(* Logix 5000 project; controller PLC_MCC1300_75F1 vendor 1 type 14 code 166 rev 32.11; software revision 32.04; part 63 of 83 *)
(* tags used below, declared in another part *)
   AUX_xInitialize : BOOL;
   CONST_rgdDestMask : DINT[32];   // Destination Mask
   CONST_tPlant : UDT_PLANT_CONSTANTS;
   GP_TrackingGetFirstPlateInConveyor : GP_TrackingGetFirstPlateInConveyor;
   GP_TrackingPresencePlate : GP_TrackingPresencePlate;
   GP_TrackingSearchPlate : GP_TrackingSearchPlate;
   M315_M1_DR_R1 : AXIS_CIP_DRIVE;
   M315_xReqStopPrevConvForPos : BOOL;
   M315Popup : MAC_Popup_ZC[2];
   M315Popup_xDrivePosEnable : BOOL;
   TMP_d : DINT;
   TMP_dIndex : DINT;
   TMP_dIndex2 : DINT;
   TMP_dIndex3 : DINT;
   TMP_dStart0 : DINT;
   TMP_dStart1 : DINT;
   TMP_dStartSearchStop : DINT;
   TMP_dStop0 : DINT;
   TMP_dStop1 : DINT;
   TMP_dStopSearchStop : DINT;
   TMP_StartPlusLength : DINT;
   TMP_xAllLiteToCullet : BOOL;
   TMP_xAtLeastOneForSideLeg : BOOL;
   TMP_xPosHead : BOOL;
   TMP_xReqStopM315M1 : BOOL;
   TMP_xReqStopM315M2 : BOOL;
   TMP_xReqStopM315M3 : BOOL;
   xAlwaysOFF : BOOL;
   xDebugOFF : BOOL;
   Z300_BufferPlate : UDT_LINE_BUFFER_PLATE;
   Z300_Conveyor : UDT_StandConv[29];
   Z300_Conveyor_IN_MOTION : MAC_Conveyor_ZC_IN_MOTION[29];
   Z300_LineTracking : UDT_LINE_TRACKING;
(* MainProgram, continued *)

   37: XIC(Z300_Conveyor[26].OUTPUT_xPositioning.0)[[XIC(Z300_Conveyor_IN_MOTION[26].DR_MAM_M[0].PC) ,XIC(xAlwaysOFF) ADD(Z300_LineTracking.rgtTrkConv[26].dStartPosition_cmm,Z300_Conveyor[26].AUX_rgdTarget_cmm[0],TMP_d) SUB(TMP_d,Z300_LineTracking.rgtTrkConv[26].dActualRamp_cmm[0],TMP_d) GEQ(Z300_BufferPlate.rgtPlate[TMP_dIndex].tTracking.dPositionHead_cmm,TMP_d) ] ,XIO(xDebugOFF) XIC(Z300_Conveyor[26].ST_xPositionReached) ][OTE(Z300_Conveyor[26].ST_xPositionReached) ,MOV(M315Popup[0].AUX_dIndexPositioning,TMP_dIndex) JSR(sbrTrackingPositioningDone,3,TMP_dIndex,TMP_xPosHead,Z300_Conveyor[26].AUX_rgdTarget_cmm[0]) ];
   38: XIC(Z300_Conveyor[27].OUTPUT_xPositioning.0)[[XIC(Z300_Conveyor_IN_MOTION[27].DR_MAM_M[0].PC) ,XIC(xAlwaysOFF) ADD(Z300_LineTracking.rgtTrkConv[26].dStartPosition_cmm,Z300_Conveyor[26].AUX_rgdTarget_cmm[0],TMP_d) SUB(TMP_d,Z300_LineTracking.rgtTrkConv[26].dActualRamp_cmm[0],TMP_d) GEQ(Z300_BufferPlate.rgtPlate[TMP_dIndex].tTracking.dPositionHead_cmm,TMP_d) ] ,XIO(xDebugOFF) XIC(Z300_Conveyor[27].ST_xPositionReached) ][OTE(Z300_Conveyor[27].ST_xPositionReached) ,MOV(M315Popup[0].AUX_dIndexPositioning,TMP_dIndex) JSR(sbrTrackingPositioningDone,3,TMP_dIndex,TMP_xPosHead,Z300_Conveyor[26].AUX_rgdTarget_cmm[0]) ];
   39: XIC(Z300_Conveyor[28].OUTPUT_xPositioning.0)[XIC(Z300_Conveyor_IN_MOTION[28].DR_MAM_M[0].PC) ,XIC(xAlwaysOFF) ADD(Z300_LineTracking.rgtTrkConv[26].dStartPosition_cmm,Z300_Conveyor[26].AUX_rgdTarget_cmm[0],TMP_d) SUB(TMP_d,Z300_LineTracking.rgtTrkConv[26].dActualRamp_cmm[0],TMP_d) GEQ(Z300_BufferPlate.rgtPlate[TMP_dIndex].tTracking.dPositionHead_cmm,TMP_d) ,XIO(xAlwaysOFF) XIC(Z300_Conveyor[28].ST_xPositionReached) ][OTE(Z300_Conveyor[28].ST_xPositionReached) ,MOV(M315Popup[0].AUX_dIndexPositioning,TMP_dIndex) JSR(sbrTrackingPositioningDone,3,TMP_dIndex,TMP_xPosHead,Z300_Conveyor[26].AUX_rgdTarget_cmm[0]) ];
   // Head positioning done
   40: [XIC(Z300_Conveyor[26].xReqPositioningHead) ,XIC(Z300_Conveyor[27].xReqPositioningHead) ,XIC(Z300_Conveyor[28].xReqPositioningHead) ][XIC(Z300_Conveyor[26].ST_xPositionReached) XIC(Z300_Conveyor[27].ST_xPositionReached) [XIC(Z300_Conveyor[28].ST_xPositionReached) ,XIO(Z300_Conveyor[28].xReqPositioningHead) ] ,XIC(Z300_Conveyor[26].xReqStop) XIO(Z300_Conveyor[26].ST_xRotationFeedback) XIC(Z300_Conveyor[27].xReqStop) XIO(Z300_Conveyor[27].ST_xRotationFeedback) [XIC(Z300_Conveyor[28].xReqStop) XIO(Z300_Conveyor[28].ST_xRotationFeedback) ,XIO(Z300_Conveyor[28].xReqPositioningHead) ] ,XIC(M315Popup[0].OS_xTimeoutPositioning) ,XIC(xDebugOFF) XIO(M315Popup[0].ST_xIndexConsPositioning) ,XIC(Z300_Conveyor[26].ST_xCleaningEnabled) ,XIC(Z300_Conveyor[26].ST_xFaulted) ,XIC(Z300_Conveyor[27].ST_xFaulted) ,XIC(Z300_Conveyor[28].ST_xFaulted) ][OTU(Z300_Conveyor[26].xReqPositioningHead) ,OTU(Z300_Conveyor[27].xReqPositioningHead) ,OTU(Z300_Conveyor[28].xReqPositioningHead) ,XIO(Z300_Conveyor[26].ST_xFaulted) XIO(Z300_Conveyor[27].ST_xFaulted) XIO(Z300_Conveyor[28].ST_xFaulted) XIO(Z300_Conveyor[26].ST_xCleaningEnabled) XIO(M315Popup[0].OS_xTimeoutPositioning) XIC(M315Popup[0].ST_xIndexConsPositioning) MOV(M315Popup[0].AUX_dIndexPositioning,TMP_dIndex) [OTL(Z300_BufferPlate.rgtPlate[TMP_dIndex].tData.tFlag.tConveyor.xDoneHeadPositioning) ,JSR(sbrTrackingPositioningDone,3,TMP_dIndex,TMP_xPosHead,Z300_Conveyor[26].AUX_rgdTarget_cmm[0]) ,MOV(M315Popup[0].AUX_dIndexPositioning,M315Popup[0].AUX_dIndexPlatePositioned) ] ,MOV(0,M315Popup[0].AUX_dIndexHead) ];
   // When plate tail has passed previous conveyor remove positioning
   41: [XIC(Z300_Conveyor[26].xReqPositioningHead) ,XIC(Z300_Conveyor[27].xReqPositioningHead) ,XIC(Z300_Conveyor[28].xReqPositioningHead) ][XIO(M315Popup[0].ST_xPrevConvFreeAfterPos) NEQ(M315Popup[0].AUX_dIndexPositioning,0) ,XIC(M315Popup[0].ST_xPrevConvFreeAfterPos) EQU(M315Popup[0].AUX_dIndexPositioning,M315Popup[0].AUX_dLastIndexFreeForPos) ][XIC(Z300_Conveyor[25].xReqPositioningHead) MOV(M315Popup[0].AUX_dIndexPositioning,TMP_dIndex) GEQ(Z300_BufferPlate.rgtPlate[TMP_dIndex].tTracking.dPositionTail_cmm,Z300_LineTracking.rgtTrkConv[25].dEndPosition_cmm) ,XIC(M315Popup[0].ST_xPrevConvFreeAfterPos) ][OTU(Z300_Conveyor[25].xReqPositioningHead) ,[XIC(Z300_Conveyor[26].ST_xRotationFeedback) ,XIC(Z300_Conveyor[26].ST_xDriveInDec) ] OTE(M315Popup[0].ST_xPrevConvFreeAfterPos) ,ONS(M315Popup[0].OS_xLastFreeForPos) MOV(M315Popup[0].AUX_dIndexPositioning,M315Popup[0].AUX_dLastIndexFreeForPos) ];
   // Tail positioning done
   42: [XIC(Z300_Conveyor[26].xReqPositioningTail) ,XIC(Z300_Conveyor[27].xReqPositioningTail) ,XIC(Z300_Conveyor[28].xReqPositioningTail) ][XIC(Z300_Conveyor[26].ST_xPositionReached) XIC(Z300_Conveyor[27].ST_xPositionReached) [XIC(Z300_Conveyor[28].ST_xPositionReached) ,XIO(Z300_Conveyor[28].xReqPositioningTail) ] ,XIC(M315Popup[0].OS_xTimeoutPositioning) ,XIO(M315Popup[0].ST_xIndexConsPositioning) ,XIC(Z300_Conveyor[26].ST_xCleaningEnabled) ,XIC(Z300_Conveyor[26].ST_xFaulted) ,XIC(Z300_Conveyor[27].ST_xFaulted) ,XIC(Z300_Conveyor[28].ST_xFaulted) ][OTU(Z300_Conveyor[26].xReqPositioningTail) ,OTU(Z300_Conveyor[27].xReqPositioningTail) ,OTU(Z300_Conveyor[28].xReqPositioningTail) ,XIO(Z300_Conveyor[26].ST_xFaulted) XIO(Z300_Conveyor[27].ST_xFaulted) XIO(Z300_Conveyor[28].ST_xFaulted) XIO(Z300_Conveyor[26].ST_xCleaningEnabled) XIO(M315Popup[0].OS_xTimeoutPositioning) MOV(M315Popup[0].AUX_tSearchPlateData.dIndex,TMP_dIndex) [OTL(Z300_BufferPlate.rgtPlate[TMP_dIndex].tData.tFlag.tConveyor.xDoneTailPositioning) ,JSR(sbrTrackingPositioningDone,3,TMP_dIndex,TMP_xPosHead,Z300_Conveyor[26].AUX_rgdTarget_cmm[0]) ,XIO(xDebugOFF) MOV(M315Popup[0].AUX_dIndexPositioning,M315Popup[0].AUX_dIndexPlatePositioned) ] ,MOV(0,M315Popup[0].AUX_dIndexTail) ];
   // Timeout positioning
   43: [[XIC(Z300_Conveyor[26].xReqPositioningHead) ,XIC(Z300_Conveyor[27].xReqPositioningHead) ,XIC(Z300_Conveyor[28].xReqPositioningHead) ] MOV(M315Popup[0].AUX_dIndexPositioning,TMP_dIndex) GEQ(Z300_BufferPlate.rgtPlate[TMP_dIndex].tTracking.dPositionHead_cmm,M315Popup[0].AUX_dPosTimeout) XIO(Z300_BufferPlate.rgtPlate[TMP_dIndex].tData.tFlag.tConveyor.xDoneHeadPositioning) ,[XIC(Z300_Conveyor[26].xReqPositioningTail) ,XIC(Z300_Conveyor[27].xReqPositioningTail) ,XIC(Z300_Conveyor[28].xReqPositioningTail) ] MOV(M315Popup[0].AUX_dIndexPositioning,TMP_dIndex) GEQ(Z300_BufferPlate.rgtPlate[TMP_dIndex].tTracking.dPositionTail_cmm,M315Popup[0].AUX_dPosTimeout) XIO(Z300_BufferPlate.rgtPlate[TMP_dIndex].tData.tFlag.tConveyor.xDoneTailPositioning) ]OTE(M315Popup[0].OS_xTimeoutPositioning);
   44: XIC(Z300_Conveyor[25].xReqPositioningHead)XIO(M315Popup[0].AUX_tSearchPlateData.xPlateHooked)OTU(Z300_Conveyor[25].xReqPositioningHead);
   45: XIC(Z300_Conveyor[25].xReqPositioningTail)XIO(M315Popup[0].AUX_tSearchPlateData.xPlateHooked)OTU(Z300_Conveyor[25].xReqPositioningTail);
   46: XIC(Z300_Conveyor[26].xReqPositioningHead)XIO(M315Popup[0].AUX_tSearchPlateData.xPlateHooked)OTU(Z300_Conveyor[26].xReqPositioningHead);
   47: XIC(Z300_Conveyor[26].xReqPositioningTail)XIO(M315Popup[0].AUX_tSearchPlateData.xPlateHooked)OTU(Z300_Conveyor[26].xReqPositioningTail);
   48: XIC(Z300_Conveyor[27].xReqPositioningHead)XIO(M315Popup[0].AUX_tSearchPlateData.xPlateHooked)OTU(Z300_Conveyor[27].xReqPositioningHead);
   49: XIC(Z300_Conveyor[27].xReqPositioningTail)XIO(M315Popup[0].AUX_tSearchPlateData.xPlateHooked)OTU(Z300_Conveyor[27].xReqPositioningTail);
   50: XIC(Z300_Conveyor[28].xReqPositioningHead)XIO(M315Popup[0].AUX_tSearchPlateData.xPlateHooked)OTU(Z300_Conveyor[28].xReqPositioningHead);
   51: XIC(Z300_Conveyor[28].xReqPositioningTail)XIO(M315Popup[0].AUX_tSearchPlateData.xPlateHooked)OTU(Z300_Conveyor[28].xReqPositioningTail);
   // #####_PRESENCE_PLATE_ON_POPUP_AFTER_POSITIONING_#####
   52: NOP();
   // Search on whole popup size
   53: ADD(0,M315Popup[0].AUX_dStartPosition_cmm,TMP_dStartSearchStop)ADD(70000,M315Popup[1].AUX_dEndPosition_cmm,TMP_dStopSearchStop)XIC(M315Popup[0].ST_xPlateToSinglePositioning)ADD(0,M315Popup[0].AUX_dStartPosition_cmm,TMP_dStartSearchStop)ADD(70000,M315Popup[0].AUX_dEndPosition_cmm,TMP_dStopSearchStop);
   54: GP_TrackingSearchPlate(GP_TrackingSearchPlate,TMP_dStopSearchStop,TMP_dStartSearchStop,0,Z300_LineTracking,M315Popup[0].tSearchPlateStop,CONST_tPlant.dNumOfConveyors,CONST_tPlant.dNumCapsConveyor,Z300_BufferPlate);
   55: XIC(M315Popup[0].tSearchPlateStop.xHeadPresence)MOV(M315Popup[0].tSearchPlateStop.rgdHeadPointer[0],M315Popup[0].AUX_dIndexPlateStop);
   56: XIO(M315Popup[0].tSearchPlateStop.xHeadPresence)XIC(M315Popup[0].tSearchPlateStop.xTailPresence)MOV(M315Popup[0].tSearchPlateStop.rgdTailPointer[0],M315Popup[0].AUX_dIndexPlateStop);
   57: [XIO(M315Popup[0].tSearchPlateStop.xHeadPresence) XIO(M315Popup[0].tSearchPlateStop.xTailPresence) ,XIC(Z300_Conveyor[26].ST_xCleaningEnabled) ]MOV(0,M315Popup[0].AUX_dIndexPlateStop);
   58: [XIC(M315Popup[0].tSearchPlateStop.xHeadPresence) ,XIC(M315Popup[0].tSearchPlateStop.xTailPresence) ][OTU(TMP_xAtLeastOneForSideLeg) ,OTL(TMP_xAllLiteToCullet) ];
   59: [XIC(M315Popup[0].tSearchPlateStop.xHeadPresence) ,XIC(M315Popup[0].tSearchPlateStop.xTailPresence) ]JSR(sbrCheckConvoyZCDestination,5,M315Popup[0].AUX_dIndexPlateStop,M315Popup[0].AUX_dDestMaskOppOpSide,CONST_rgdDestMask[24],TMP_xAtLeastOneForSideLeg,TMP_xAllLiteToCullet,TMP_xAtLeastOneForSideLeg,TMP_xAllLiteToCullet)XIC(TMP_xAtLeastOneForSideLeg)[EQU(M315Popup[0].AUX_dIndexPositioning,M315Popup[0].AUX_dIndexPlateStop) ,EQU(M315Popup[0].AUX_dIndexPlatePositioned,M315Popup[0].AUX_dIndexPlateStop) ,EQU(M315Popup[0].tSearchPlateStop.rgdHeadPointer[1],M315Popup[0].AUX_dIndexPlateStop) ,EQU(M315Popup[0].tSearchPlateStop.rgdHeadPointer[1],M315Popup[0].AUX_dIndexPlatePositioned) ,EQU(M315Popup[0].tSearchPlateStop.rgdTailPointer[1],M315Popup[0].AUX_dIndexPlateStop) ,EQU(M315Popup[0].tSearchPlateStop.rgdTailPointer[1],M315Popup[0].AUX_dIndexPlatePositioned) ,XIO(xDebugOFF) ]OTE(M315Popup[0].ST_xPlateStopToPopup);
   // IndexPlatePositioned valorizzata qui solo per la simulazione (da togliere)
   60: XIC(M315Popup[0].AUX_tSearchPlateData.xPlateHooked)[XIC(M315Popup[0].tSearchPlateStop.xHeadPresence) ,XIC(M315Popup[0].tSearchPlateStop.xTailPresence) ,XIO(M315Popup[1].ST_xPlateToSinglePositioning) EQU(M315Popup[0].AUX_dIndexPositioning,Z300_LineTracking.rgtTrkConv[26].Cap[0].dPointer) ,XIO(M315Popup[1].ST_xPlateToSinglePositioning) EQU(M315Popup[0].AUX_dIndexPlatePositioned,Z300_LineTracking.rgtTrkConv[26].Cap[0].dPointer) ][XIC(TMP_xPosHead) MOV(M315Popup[0].AUX_dIndexPositioning,TMP_dIndex) XIC(Z300_BufferPlate.rgtPlate[TMP_dIndex].tData.tFlag.tConveyor.xDoneHeadPositioning) ,XIO(TMP_xPosHead) MOV(M315Popup[0].AUX_dIndexPositioning,TMP_dIndex) XIC(Z300_BufferPlate.rgtPlate[TMP_dIndex].tData.tFlag.tConveyor.xDoneTailPositioning) ]XIO(M315Popup_xDrivePosEnable)XIC(M315Popup[0].ST_xPlateStopToPopup)[OTE(TMP_xReqStopM315M1) ,OTE(TMP_xReqStopM315M2) ,XIO(M315Popup[0].ST_xPlateToSinglePositioning) OTE(TMP_xReqStopM315M3) ];
   61: XIO(xDebugOFF)XIC(Z300_Conveyor[26].OUTPUT_xPositioning.0)OTE(Z300_Conveyor[26].xReqBypassEndStop);
   62: XIO(xDebugOFF)XIC(Z300_Conveyor[27].OUTPUT_xPositioning.0)OTE(Z300_Conveyor[27].xReqBypassEndStop);
   63: XIO(xDebugOFF)XIC(Z300_Conveyor[28].OUTPUT_xPositioning.0)OTE(Z300_Conveyor[28].xReqBypassEndStop);
   64: [XIC(TMP_xReqStopM315M1) ,XIC(M315Popup[0].PH_xDescend) ]OTE(Z300_Conveyor[26].xReqStop);
   65: [XIC(TMP_xReqStopM315M2) ,XIC(M315Popup[0].PH_xDescend) ]OTE(Z300_Conveyor[27].xReqStop);
   66: [XIC(TMP_xReqStopM315M3) ,XIC(M315Popup[1].PH_xDescend) ]OTE(Z300_Conveyor[28].xReqStop);
   // Stop tracking update while ending positioning
   67: XIO(xDebugOFF)XIC(M315Popup[0].AUX_tSearchPlateData.xPlateHooked)MOV(M315Popup[0].AUX_dIndexPositioning,TMP_dIndex)XIC(M315Popup_xDrivePosEnable)[ADD(Z300_LineTracking.rgtTrkConv[26].dStartPosition_cmm,Z300_Conveyor[26].AUX_rgdTarget_cmm[0],TMP_d) SUB(TMP_d,Z300_LineTracking.rgtTrkConv[26].dActualRamp_cmm[0],TMP_d) GEQ(Z300_BufferPlate.rgtPlate[TMP_dIndex].tTracking.dPositionHead_cmm,TMP_d) ,ADD(Z300_LineTracking.rgtTrkConv[26].dStartPosition_cmm,Z300_BufferPlate.rgtPlate[TMP_dIndex].tData.rgtCap[0].dConvTotLength_cmm,TMP_StartPlusLength) GEQ(Z300_BufferPlate.rgtPlate[TMP_dIndex].tTracking.dPositionHead_cmm,TMP_StartPlusLength) ][XIC(M315Popup[0].ST_xPlateStopToPopup) ,XIC(M315Popup[1].ST_xPlateStopToPopup) ]XIC(Z300_Conveyor_IN_MOTION[26].DR_MAM_M[0].IP)XIO(Z300_Conveyor_IN_MOTION[26].DR_MAM_M[0].PC)XIO(Z300_Conveyor_IN_MOTION[26].DR_MAM_M[0].ER)[OTE(Z300_BufferPlate.rgtPlate[TMP_dIndex].tTracking.xHoldAdvancement) ,ADD(M315Popup[0].AUX_dPosPhotocell_cmm,Z300_Conveyor[26].AUX_rgdTarget_cmm[0],TMP_d) JSR(sbrUpdateTrackingConvoyPosition,2,TMP_dIndex,TMP_d) ];
   // Stop tracking update while ending positioning
   68: XIC(M315Popup[0].AUX_tSearchPlateData.xPlateHooked)[XIC(Z300_LineTracking.rgtTrkConv[26].xGlassPresence) ,XIC(Z300_LineTracking.rgtTrkConv[27].xGlassPresence) ,XIC(Z300_LineTracking.rgtTrkConv[28].xGlassPresence) ]MOV(M315Popup[0].AUX_dIndexPositioning,TMP_dIndex)[LES(Z300_BufferPlate.rgtPlate[TMP_dIndex].tData.dTotalCaps,2) ,XIO(xDebugOFF) ]XIC(M315Popup_xDrivePosEnable)XIO(M315_M1_DR_R1.Registration1InputStatus)[ADD(Z300_LineTracking.rgtTrkConv[26].dStartPosition_cmm,Z300_Conveyor[26].AUX_rgdTarget_cmm[0],TMP_d) SUB(TMP_d,Z300_LineTracking.rgtTrkConv[26].dActualRamp_cmm[0],TMP_d) GEQ(Z300_BufferPlate.rgtPlate[TMP_dIndex].tTracking.dPositionHead_cmm,TMP_d) ,ADD(Z300_LineTracking.rgtTrkConv[26].dStartPosition_cmm,Z300_BufferPlate.rgtPlate[TMP_dIndex].tData.rgtCap[0].dConvTotLength_cmm,TMP_StartPlusLength) GEQ(Z300_BufferPlate.rgtPlate[TMP_dIndex].tTracking.dPositionHead_cmm,TMP_StartPlusLength) ]OTE(M315_xReqStopPrevConvForPos);
   69: XIO(xDebugOFF)XIC(Z300_BufferPlate.rgtPlate[TMP_dIndex].tTracking.xHoldAdvancement)GRT(Z300_BufferPlate.rgtPlate[TMP_dIndex].tTracking.dNextCapIndex,0)MOV(Z300_BufferPlate.rgtPlate[TMP_dIndex].tTracking.dNextCapIndex,TMP_dIndex2)OTE(Z300_BufferPlate.rgtPlate[TMP_dIndex2].tTracking.xHoldAdvancement);
   70: XIO(xDebugOFF)XIC(Z300_BufferPlate.rgtPlate[TMP_dIndex2].tTracking.xHoldAdvancement)GRT(Z300_BufferPlate.rgtPlate[TMP_dIndex2].tTracking.dNextCapIndex,0)MOV(Z300_BufferPlate.rgtPlate[TMP_dIndex2].tTracking.dNextCapIndex,TMP_dIndex3)OTE(Z300_BufferPlate.rgtPlate[TMP_dIndex3].tTracking.xHoldAdvancement);
   // #####_PRESENCE_PLATE_UNDER_POPUP_#####
   71: NOP();
   72: [XIC(Z300_Conveyor[25].ST_xRotationFeedback) SUB(M315Popup[0].AUX_dStartPosition_cmm,25000,TMP_dStart0) ,XIO(Z300_Conveyor[25].ST_xRotationFeedback) SUB(M315Popup[0].AUX_dStartPosition_cmm,0,TMP_dStart0) ]ADD(M315Popup[0].AUX_dEndPosition_cmm,70000,TMP_dStop0)[XIC(Z300_Conveyor[25].ST_xRotationFeedback) SUB(M315Popup[1].AUX_dStartPosition_cmm,75000,TMP_dStart1) ,XIO(Z300_Conveyor[25].ST_xRotationFeedback) SUB(M315Popup[1].AUX_dStartPosition_cmm,25000,TMP_dStart1) ]ADD(M315Popup[1].AUX_dEndPosition_cmm,55000,TMP_dStop1)GP_TrackingPresencePlate(GP_TrackingPresencePlate,TMP_dStart0,TMP_dStop0,0,Z300_LineTracking,M315Popup[0].ST_xPlateUnderPopup)GP_TrackingPresencePlate(GP_TrackingPresencePlate,TMP_dStart1,TMP_dStop1,0,Z300_LineTracking,M315Popup[1].ST_xPlateUnderPopup);
   73: XIC(M315Popup[0].AUX_tSearchPlateData.xPlateHooked)GRT(M315Popup[0].AUX_dIndexPositioning,0)MOV(M315Popup[0].AUX_dIndexPositioning,TMP_dIndex)[XIC(TMP_xPosHead) GEQ(Z300_BufferPlate.rgtPlate[TMP_dIndex].tTracking.dPositionHead_cmm,M315Popup[0].AUX_tSearchPlateData.dPositionStopHooked_cmm) ,XIO(TMP_xPosHead) GEQ(Z300_BufferPlate.rgtPlate[TMP_dIndex].tTracking.dPositionTail_cmm,M315Popup[0].AUX_tSearchPlateData.dPositionStopHooked_cmm) ][OSR(M315Popup[0].AUX_tSearchPlateData.OSR_xPlateOutHooked,M315Popup[0].AUX_tSearchPlateData.OS_xPlateOutHooked) ,OTE(M315Popup[0].ST_xPopupChangeDest) ];
   // #####_Change_Destination_#####
   74: XIC(M315Popup[0].ST_xPopupChangeDest)[JSR(sbrRedestConvoyCapZC,5,M315Popup[0].AUX_dIndexPositioning,M315Popup[0].AUX_dDestMaskOppOpSide,0,1,CONST_rgdDestMask[24]) ,OTU(M315Popup[0].AUX_tSearchPlateData.xPlateHooked) ,MOV(0,M315Popup[0].AUX_dIndexPositioning) ,MOV(0,M315Popup[0].AUX_dIndexPlatePositioned) ];
   75: [XIC(M315Popup[0].AUX_tSearchPlateData.OS_xPlateOutHooked) ,XIC(M315Popup[0].AUX_tSearchPlateData.xPlateHooked) XIO(M315Popup[0].AUX_tSearchPlateData.xIndexCons) ,XIC(Z300_Conveyor[26].ST_xCleaningEnabled) ][MOV(0,M315Popup[0].AUX_dIndexPositioning) ,OTU(M315Popup[0].AUX_tSearchPlateData.xPlateHooked) ,OTU(Z300_Conveyor[26].xReqPositioningHead) ,OTU(Z300_Conveyor[27].xReqPositioningHead) ,OTU(Z300_Conveyor[28].xReqPositioningHead) ,OTU(Z300_Conveyor[26].xReqPositioningTail) ,OTU(Z300_Conveyor[27].xReqPositioningTail) ,OTU(Z300_Conveyor[28].xReqPositioningTail) ];
   // Check if there is a cap destined to popup during a restart of the CPU and make redestination (second conveyor)
   76: XIC(AUX_xInitialize)XIC(M315Popup[1].ST_xPlateStopToPopup)GP_TrackingGetFirstPlateInConveyor(GP_TrackingGetFirstPlateInConveyor,Z300_LineTracking.rgtTrkConv[28],CONST_tPlant.dNumCapsConveyor,GP_TrackingGetFirstPlateInConveyor.OUT_dIndex,GP_TrackingGetFirstPlateInConveyor.OUT_dHeadPos)GRT(GP_TrackingGetFirstPlateInConveyor.OUT_dIndex,0)GRT(GP_TrackingGetFirstPlateInConveyor.OUT_dHeadPos,M315Popup[1].AUX_dStartPosition_cmm)LES(GP_TrackingGetFirstPlateInConveyor.OUT_dHeadPos,M315Popup[1].AUX_dEndPosition_cmm)MOV(GP_TrackingGetFirstPlateInConveyor.OUT_dIndex,M315Popup[0].AUX_dIndexPlatePositioned)OTE(M315Popup[1].OS_xChangeDestAfterRestart);
   // Change destination aftet restart (second conveyor)
   77: XIC(M315Popup[1].OS_xChangeDestAfterRestart)[JSR(sbrRedestConvoyCapZC,5,M315Popup[0].AUX_dIndexPlatePositioned,M315Popup[0].AUX_dDestMaskOppOpSide,0,1,CONST_rgdDestMask[24]) ,JSR(sbrTrackingIndexTailConvoy,1,M315Popup[0].AUX_dIndexPlatePositioned,M315Popup[0].AUX_dIndexPlateFree) ,OTU(M315Popup[0].AUX_tSearchPlateData.xPlateHooked) ,MOV(0,M315Popup[0].AUX_dIndexPositioning) ,MOV(0,M315Popup[0].AUX_dIndexPlatePositioned) ];
   // Check if there is a cap destined to popup during a restart of the CPU and make redestination (first conveyor)
   78: XIC(AUX_xInitialize)XIC(M315Popup[0].ST_xPlateStopToPopup)GP_TrackingGetFirstPlateInConveyor(GP_TrackingGetFirstPlateInConveyor,Z300_LineTracking.rgtTrkConv[22],CONST_tPlant.dNumCapsConveyor,GP_TrackingGetFirstPlateInConveyor.OUT_dIndex,GP_TrackingGetFirstPlateInConveyor.OUT_dHeadPos)GRT(GP_TrackingGetFirstPlateInConveyor.OUT_dIndex,0)GRT(GP_TrackingGetFirstPlateInConveyor.OUT_dHeadPos,M315Popup[0].AUX_dStartPosition_cmm)LES(GP_TrackingGetFirstPlateInConveyor.OUT_dHeadPos,M315Popup[0].AUX_dEndPosition_cmm)MOV(GP_TrackingGetFirstPlateInConveyor.OUT_dIndex,M315Popup[0].AUX_dIndexPlatePositioned)OTE(M315Popup[0].OS_xChangeDestAfterRestart);
   // Change destination aftet restart (first conveyor)
   79: XIC(M315Popup[0].OS_xChangeDestAfterRestart)[JSR(sbrRedestConvoyCapZC,5,M315Popup[0].AUX_dIndexPlatePositioned,M315Popup[0].AUX_dDestMaskOppOpSide,0,1,CONST_rgdDestMask[24]) ,JSR(sbrTrackingIndexTailConvoy,1,M315Popup[0].AUX_dIndexPlatePositioned,M315Popup[0].AUX_dIndexPlateFree) ,OTU(M315Popup[0].AUX_tSearchPlateData.xPlateHooked) ,MOV(0,M315Popup[0].AUX_dIndexPositioning) ,MOV(0,M315Popup[0].AUX_dIndexPlatePositioned) ];
   80: NOP();
   // #####_Lifting_#####
   81: NOP();
   // Plate in position to raise
   82: XIO(Z300_Conveyor[23].ST_xCleaningEnabled)[XIC(M315Popup[0].AUX_tSearchPlateData.xPlateHooked) GRT(M315Popup[0].AUX_dIndexPositioning,0) MOV(M315Popup[0].AUX_dIndexPositioning,TMP_dIndex) [XIC(TMP_xPosHead) XIC(Z300_BufferPlate.rgtPlate[TMP_dIndex].tData.tFlag.tConveyor.xDoneHeadPositioning) ,XIO(TMP_xPosHead) XIC(Z300_BufferPlate.rgtPlate[TMP_dIndex].tData.tFlag.tConveyor.xDoneTailPositioning) ] ,XIC(M315Popup[0].ST_xPlateInPositionToRise) ]XIC(M315Popup[0].ST_xPlateStopToPopup)[XIC(Z300_Conveyor[26].xReqStop) XIO(Z300_Conveyor[26].INPUT_xDriveDeceleration.0) XIO(Z300_Conveyor[26].INPUT_xDriveFeedback.0) ,XIC(Z300_Conveyor[27].xReqStop) XIO(Z300_Conveyor[27].INPUT_xDriveDeceleration.0) XIO(Z300_Conveyor[27].INPUT_xDriveFeedback.0) ,XIC(Z300_Conveyor[28].xReqStop) XIO(Z300_Conveyor[28].INPUT_xDriveDeceleration.0) XIO(Z300_Conveyor[28].INPUT_xDriveFeedback.0) ]XIO(M315Popup[0].ST_xRequestRise)XIO(M315Popup[1].ST_xRequestRise)[OTE(M315Popup[0].ST_xPlateInPositionToRise) ,EQU(M315Popup[0].AUX_dIndexPlatePositioned,0) MOV(M315Popup[0].AUX_dIndexPositioning,M315Popup[0].AUX_dIndexPlatePositioned) ];
